screen "RIO 02 Digital Inputs" 1280x800, template "Template"
   on GenerateScreen: "TitleUpdater"()
   TextField "Text field_37" at 16,52 size 476x26; Text 'RIO #2 (Remote Inputs & Outputs Panel No. 2)'
   TextField "Text field_38" at 16,122 size 55x22; Text 'I15.0'
   TextField "Text field_39" at 16,157 size 55x22; Text 'I15.1'
   TextField "Text field_40" at 16,193 size 55x22; Text 'I15.2'
   TextField "Text field_41" at 16,229 size 55x22; Text 'I15.3'
   TextField "Text field_42" at 16,265 size 55x22; Text 'I15.4'
   TextField "Text field_43" at 16,301 size 55x22; Text 'I15.5'
   TextField "Text field_44" at 16,337 size 55x22; Text 'I15.6'
   TextField "Text field_45" at 16,373 size 55x22; Text 'I15.7'
   Circle "Circle_33" at 76,123 size 20x20
      Appearance <- "Tank 2P GTT Isolation Valve Feedback - Opened"
   Circle "Circle_34" at 76,158 size 20x20
      Appearance <- "Tank 2P GTT Isolation Valve Feedback - Closed"
   Circle "Circle_35" at 76,194 size 20x20
      Appearance <- "Tank 2P Tank Vent Valve 1 Feedback - Opened"
   Circle "Circle_36" at 76,230 size 20x20
      Appearance <- "Tank 2P Tank Vent Valve 1 Feedback - Closed"
   Circle "Circle_37" at 76,265 size 20x20
      Appearance <- "Tank 2P Tank Vent Valve 2 Feedback - Opened"
   Circle "Circle_38" at 76,301 size 20x20
      Appearance <- "Tank 2P Tank Vent Valve 2 Feedback - Closed"
   Circle "Circle_39" at 76,337 size 20x20
      Appearance <- "RIO2_SPR_DI_15_6"
   Circle "Circle_40" at 76,373 size 20x20
      Appearance <- "RIO2_SPR_DI_15_7"
   TextField "Text field_46" at 33,90 size 49x26; Text 'I0'
   TextField "Text field_47" at 16,441 size 55x22; Text 'I18.0'
   TextField "Text field_48" at 16,476 size 55x22; Text 'I18.1'
   TextField "Text field_49" at 16,512 size 55x22; Text 'I18.2'
   TextField "Text field_50" at 16,548 size 55x22; Text 'I18.3'
   TextField "Text field_51" at 16,584 size 55x22; Text 'I18.4'
   TextField "Text field_52" at 16,620 size 55x22; Text 'I18.5'
   TextField "Text field_53" at 16,656 size 55x22; Text 'I18.6'
   TextField "Text field_54" at 16,692 size 55x22; Text 'I18.7'
   Circle "Circle_41" at 76,442 size 20x20
      Appearance <- "Tank 2S GTT Isolation Valve Feedback - Opened"
   Circle "Circle_42" at 76,477 size 20x20
      Appearance <- "Tank 2S GTT Isolation Valve Feedback - Closed"
   Circle "Circle_43" at 76,513 size 20x20
      Appearance <- "Tank 2S Tank Vent Valve 1 Feedback - Opened"
   Circle "Circle_44" at 76,549 size 20x20
      Appearance <- "Tank 2S Tank Vent Valve 1 Feedback - Closed"
   Circle "Circle_45" at 76,585 size 20x20
      Appearance <- "Tank 2S Tank Vent Valve 2 Feedback - Opened"
   Circle "Circle_46" at 76,621 size 20x20
      Appearance <- "Tank 2S Tank Vent Valve 2 Feedback - Closed"
   Circle "Circle_47" at 76,657 size 20x20
      Appearance <- "RIO2_SPR_DI_18_6"
   Circle "Circle_48" at 76,693 size 20x20
      Appearance <- "RIO2_SPR_DI_18_7"
   TextField "Text field_55" at 33,409 size 49x26; Text 'I1'
   TextField "Text field_56" at 548,122 size 55x22; Text 'I21.0'
   TextField "Text field_57" at 548,157 size 55x22; Text 'I21.1'
   TextField "Text field_58" at 548,193 size 55x22; Text 'I21.2'
   TextField "Text field_59" at 548,229 size 55x22; Text 'I21.3'
   TextField "Text field_60" at 548,265 size 55x22; Text 'I21.4'
   TextField "Text field_61" at 548,301 size 55x22; Text 'I21.5'
   TextField "Text field_62" at 548,337 size 55x22; Text 'I21.6'
   TextField "Text field_63" at 548,373 size 55x22; Text 'I21.7'
   Circle "Circle_49" at 608,122 size 20x20
      Appearance <- "Tank 2P BWT Level High High Switch"
   Circle "Circle_50" at 608,157 size 20x20
      Appearance <- "RIO2 Tanks Pressure Switch Hi Hi"
   Circle "Circle_51" at 608,193 size 20x20
      Appearance <- "Tank 2S BWT Level High High Switch"
   Circle "Circle_52" at 608,229 size 20x20
      Appearance <- "RIO2_SPR_DI_21_3"
   Circle "Circle_53" at 608,265 size 20x20
      Appearance <- "RIO2_SPR_DI_21_4"
   Circle "Circle_54" at 608,301 size 20x20
      Appearance <- "RIO2_SPR_DI_21_5"
   Circle "Circle_55" at 608,337 size 20x20
      Appearance <- "RIO2_SPR_DI_21_6"
   Circle "Circle_56" at 608,373 size 20x20
      Appearance <- "RIO2_SPR_DI_21_7"
   TextField "Text field_64" at 570,90 size 49x26; Text 'I2'
   Button "HmiScreenItemData_1" at 1,1 size 150x43; TextOn 'Back'; TextOff 'Commissioning'
      on Release: ActivateScreen("Commissioning Main Page", 0)
   TextField "Text field_107" at 105,114 size 382x38; Text 'Tank 2P GTT Isolation Valve Feedback - Opened CV422'
   TextField "Text field_108" at 105,149 size 374x38; Text 'Tank 2P GTT Isolation Valve Feedback - Closed CV422'
   TextField "Text field_109" at 105,184 size 371x38; Text 'Tank 2P Tank Vent Valve 1 Feedback - Opened CV441-2P1'
   TextField "Text field_110" at 105,220 size 363x38; Text 'Tank 2P Tank Vent Valve 1 Feedback - Closed CV441-2P1'
   TextField "Text field_111" at 105,255 size 371x38; Text 'Tank 2P Tank Vent Valve 2 Feedback - Opened CV441-2P2'
   TextField "Text field_112" at 105,291 size 363x38; Text 'Tank 2P Tank Vent Valve 2 Feedback - Closed CV441-2P2'
   TextField "Text field_113" at 104,328 size 100x21; Text 'Spare Input'
   TextField "Text field_114" at 104,365 size 100x21; Text 'Spare Input'
   TextField "Text field_116" at 102,429 size 382x38; Text 'Tank 2S GTT Isolation Valve Feedback - Opened CV421-2S'
   TextField "Text field_117" at 102,465 size 374x38; Text 'Tank 2S GTT Isolation Valve Feedback - Closed CV421-2S'
   TextField "Text field_118" at 102,501 size 371x38; Text 'Tank 2S Tank Vent Valve 1 Feedback - Opened CV440-2SA'
   TextField "Text field_119" at 102,537 size 363x38; Text 'Tank 2S Tank Vent Valve 1 Feedback - Closed CV440-2SA'
   TextField "Text field_120" at 102,573 size 371x38; Text 'Tank 2S Tank Vent Valve 2 Feedback - Opened CV440-2SB'
   TextField "Text field_121" at 102,609 size 363x38; Text 'Tank 2S Tank Vent Valve 2 Feedback - Closed CV440-2SB'
   TextField "Text field_122" at 102,690 size 100x21; Text 'Spare Input'
   TextField "Text field_123" at 636,113 size 294x38; Text 'Tank 2P BWT Level High High Switch LS425-2P'
   TextField "Text field_124" at 636,148 size 270x38; Text 'RIO2 Tanks Pressure Switch Hi Hi PS436-2P/2S'
   TextField "Text field_125" at 636,184 size 294x38; Text 'Tank 2S BWT Level High High Switch LS422-2S'
   TextField "Text field_126" at 636,219 size 100x21; Text 'Spare Input'
   TextField "Text field_127" at 636,255 size 100x21; Text 'Spare Input'
   TextField "Text field_128" at 636,291 size 100x21; Text 'Spare Input'
   TextField "Text field_129" at 636,328 size 100x21; Text 'Spare Input'
   TextField "Text field_130" at 636,366 size 100x21; Text 'Spare Input'
   TextField "Text field_115" at 102,654 size 100x21; Text 'Spare Input'
   AlarmView "Alarm view_1" at 0,777 size 1280x23
   Group "Group" at 455,41 size 373x50
   Button "HmiScreenItemData_8" at 469,45 size 355x40; TextOn 'Back'; TextOff 'Text'
      on Click: "TitleUpdater"()
   TextField "Screen title" at 455,41 size 373x50; Text 'Screen title'

screen "RIO 03 Digital Inputs" 1280x800, template "Template"
   on GenerateScreen: "TitleUpdater"()
   TextField "Text field_37" at 16,52 size 476x26; Text 'RIO #3 (Remote Inputs & Outputs Panel No. 3)'
   TextField "Text field_38" at 16,122 size 55x22; Text 'I27.0'
   TextField "Text field_39" at 16,157 size 55x22; Text 'I27.1'
   TextField "Text field_40" at 16,193 size 55x22; Text 'I27.2'
   TextField "Text field_41" at 16,229 size 55x22; Text 'I27.3'
   TextField "Text field_42" at 16,265 size 55x22; Text 'I27.4'
   TextField "Text field_43" at 16,301 size 55x22; Text 'I27.5'
   TextField "Text field_44" at 16,337 size 55x22; Text 'I27.6'
   TextField "Text field_45" at 16,373 size 55x22; Text 'I27.7'
   Circle "Circle_33" at 76,123 size 20x20
      Appearance <- "Tank 3P GTT Isolation Valve Feedback - Opened"
   Circle "Circle_34" at 76,158 size 20x20
      Appearance <- "Tank 3P GTT Isolation Valve Feedback - Closed"
   Circle "Circle_35" at 76,194 size 20x20
      Appearance <- "Tank 3P Tank Vent Valve 1 Feedback - Opened"
   Circle "Circle_36" at 76,230 size 20x20
      Appearance <- "Tank 3P Tank Vent Valve 1 Feedback - Closed"
   Circle "Circle_37" at 76,265 size 20x20
      Appearance <- "Tank 3P Tank Vent Valve 2 Feedback - Opened"
   Circle "Circle_38" at 76,301 size 20x20
      Appearance <- "Tank 3P Tank Vent Valve 2 Feedback - Closed"
   Circle "Circle_39" at 76,337 size 20x20
      Appearance <- "RIO3_SPR_DI_27_6"
   Circle "Circle_40" at 76,373 size 20x20
      Appearance <- "RIO3_SPR_DI_27_7"
   TextField "Text field_46" at 33,90 size 49x26; Text 'I0'
   TextField "Text field_47" at 16,441 size 55x22; Text 'I30.0'
   TextField "Text field_48" at 16,476 size 55x22; Text 'I30.1'
   TextField "Text field_49" at 16,512 size 55x22; Text 'I30.2'
   TextField "Text field_50" at 16,548 size 55x22; Text 'I30.3'
   TextField "Text field_51" at 16,584 size 55x22; Text 'I30.4'
   TextField "Text field_52" at 16,620 size 55x22; Text 'I30.5'
   TextField "Text field_53" at 16,656 size 55x22; Text 'I30.6'
   TextField "Text field_54" at 16,692 size 55x22; Text 'I30.7'
   Circle "Circle_41" at 76,442 size 20x20
      Appearance <- "Tank 3S GTT Isolation Valve Feedback - Opened"
   Circle "Circle_42" at 76,477 size 20x20
      Appearance <- "Tank 3S GTT Isolation Valve Feedback - Closed"
   Circle "Circle_43" at 76,513 size 20x20
      Appearance <- "Tank 3S Tank Vent Valve 1 Feedback - Opened"
   Circle "Circle_44" at 76,549 size 20x20
      Appearance <- "Tank 3S Tank Vent Valve 1 Feedback - Closed"
   Circle "Circle_45" at 76,585 size 20x20
      Appearance <- "Tank 3S Tank Vent Valve 2 Feedback - Opened"
   Circle "Circle_46" at 76,621 size 20x20
      Appearance <- "Tank 3S Tank Vent Valve 2 Feedback - Closed"
   Circle "Circle_47" at 76,657 size 20x20
      Appearance <- "RIO3_SPR_DI_30_6"
   Circle "Circle_48" at 76,693 size 20x20
      Appearance <- "RIO3_SPR_DI_30_7"
   TextField "Text field_55" at 33,409 size 49x26; Text 'I1'
   TextField "Text field_56" at 548,122 size 55x22; Text 'I33.0'
   TextField "Text field_57" at 548,157 size 55x22; Text 'I33.1'
   TextField "Text field_58" at 548,193 size 55x22; Text 'I33.2'
   TextField "Text field_59" at 548,229 size 55x22; Text 'I33.3'
   TextField "Text field_60" at 548,265 size 55x22; Text 'I33.4'
   TextField "Text field_61" at 548,301 size 55x22; Text 'I33.5'
   TextField "Text field_62" at 548,337 size 55x22; Text 'I33.6'
   TextField "Text field_63" at 548,373 size 55x22; Text 'I33.7'
   Circle "Circle_49" at 608,122 size 20x20
      Appearance <- "Tank 3P BWT Level High High Switch"
   Circle "Circle_50" at 608,157 size 20x20
      Appearance <- "RIO3 Tanks Pressure Switch Hi Hi"
   Circle "Circle_51" at 608,193 size 20x20
      Appearance <- "Tank 3S BWT Level High High Switch"
   Circle "Circle_52" at 608,229 size 20x20
      Appearance <- "RIO3_SPR_DI_33_3"
   Circle "Circle_53" at 608,265 size 20x20
      Appearance <- "RIO3_SPR_DI_33_4"
   Circle "Circle_54" at 608,301 size 20x20
      Appearance <- "RIO3_SPR_DI_33_5"
   Circle "Circle_55" at 608,337 size 20x20
      Appearance <- "RIO3_SPR_DI_33_6"
   Circle "Circle_56" at 608,373 size 20x20
      Appearance <- "RIO3_SPR_DI_33_7"
   TextField "Text field_64" at 570,90 size 49x26; Text 'I2'
   Button "HmiScreenItemData_1" at 1,1 size 150x43; TextOn 'Back'; TextOff 'Commissioning'
      on Release: ActivateScreen("Commissioning Main Page", 0)
   TextField "Text field_107" at 105,114 size 382x38; Text 'Tank 3P GTT Isolation Valve Feedback - Opened CV422'
   TextField "Text field_108" at 105,149 size 374x38; Text 'Tank 3P GTT Isolation Valve Feedback - Closed CV422'
   TextField "Text field_109" at 105,184 size 371x38; Text 'Tank 3P Tank Vent Valve 1 Feedback - Opened CV441-3P1'
   TextField "Text field_110" at 105,220 size 363x38; Text 'Tank 3P Tank Vent Valve 1 Feedback - Closed CV441-3P1'
   TextField "Text field_111" at 105,255 size 371x38; Text 'Tank 3P Tank Vent Valve 2 Feedback - Opened CV441-3P2'
   TextField "Text field_112" at 105,291 size 363x38; Text 'Tank 3P Tank Vent Valve 2 Feedback - Closed CV441-3P2'
   TextField "Text field_113" at 104,328 size 100x21; Text 'Spare Input'
   TextField "Text field_114" at 104,365 size 100x21; Text 'Spare Input'
   TextField "Text field_116" at 102,429 size 382x38; Text 'Tank 3S GTT Isolation Valve Feedback - Opened CV421-3S'
   TextField "Text field_117" at 102,465 size 374x38; Text 'Tank 3S GTT Isolation Valve Feedback - Closed CV421-3S'
   TextField "Text field_118" at 102,501 size 371x38; Text 'Tank 3S Tank Vent Valve 1 Feedback - Opened CV440-3SA'
   TextField "Text field_119" at 102,537 size 363x38; Text 'Tank 3S Tank Vent Valve 1 Feedback - Closed CV440-3SA'
   TextField "Text field_120" at 102,573 size 371x38; Text 'Tank 3S Tank Vent Valve 2 Feedback - Opened CV440-3SB'
   TextField "Text field_121" at 102,609 size 363x38; Text 'Tank 3S Tank Vent Valve 2 Feedback - Closed CV440-3SB'
   TextField "Text field_122" at 102,690 size 100x21; Text 'Spare Input'
   TextField "Text field_123" at 636,113 size 294x38; Text 'Tank 3P BWT Level High High Switch LS425-3P'
   TextField "Text field_124" at 636,148 size 270x38; Text 'RIO3 Tanks Pressure Switch Hi Hi PS436-3P/3S'
   TextField "Text field_125" at 636,184 size 294x38; Text 'Tank 3S BWT Level High High Switch LS422-3S'
   TextField "Text field_126" at 636,219 size 100x21; Text 'Spare Input'
   TextField "Text field_127" at 636,255 size 100x21; Text 'Spare Input'
   TextField "Text field_128" at 636,291 size 100x21; Text 'Spare Input'
   TextField "Text field_129" at 636,328 size 100x21; Text 'Spare Input'
   TextField "Text field_130" at 636,366 size 100x21; Text 'Spare Input'
   TextField "Text field_115" at 102,654 size 100x21; Text 'Spare Input'
   AlarmView "Alarm view_1" at 0,777 size 1280x23
   Group "Group" at 455,41 size 373x50
   Button "HmiScreenItemData_8" at 469,45 size 355x40; TextOn 'Back'; TextOff 'Text'
      on Click: "TitleUpdater"()
   TextField "Screen title" at 455,41 size 373x50; Text 'Screen title'

screen "RIO 04 Digital Inputs" 1280x800, template "Template"
   on GenerateScreen: "TitleUpdater"()
   TextField "Text field_37" at 16,52 size 476x26; Text 'RIO #4 (Remote Inputs & Outputs Panel No. 4)'
   TextField "Text field_38" at 16,122 size 55x22; Text 'I39.0'
   TextField "Text field_39" at 16,157 size 55x22; Text 'I39.1'
   TextField "Text field_40" at 16,193 size 55x22; Text 'I39.2'
   TextField "Text field_41" at 16,229 size 55x22; Text 'I39.3'
   TextField "Text field_42" at 16,265 size 55x22; Text 'I39.4'
   TextField "Text field_43" at 16,301 size 55x22; Text 'I39.5'
   TextField "Text field_44" at 16,337 size 55x22; Text 'I39.6'
   TextField "Text field_45" at 16,373 size 55x22; Text 'I39.7'
   Circle "Circle_33" at 76,123 size 20x20
      Appearance <- "Tank 4P GTT Isolation Valve Feedback - Opened"
   Circle "Circle_34" at 76,158 size 20x20
      Appearance <- "Tank 4P GTT Isolation Valve Feedback - Closed"
   Circle "Circle_35" at 76,194 size 20x20
      Appearance <- "Tank 4P Tank Vent Valve 1 Feedback - Opened"
   Circle "Circle_36" at 76,230 size 20x20
      Appearance <- "Tank 4P Tank Vent Valve 1 Feedback - Closed"
   Circle "Circle_37" at 76,265 size 20x20
      Appearance <- "Tank 4P Tank Vent Valve 2 Feedback - Opened"
   Circle "Circle_38" at 76,301 size 20x20
      Appearance <- "Tank 4P Tank Vent Valve 2 Feedback - Closed"
   Circle "Circle_39" at 76,337 size 20x20
      Appearance <- "RIO4_SPR_DI_139_6"
   Circle "Circle_40" at 76,373 size 20x20
      Appearance <- "RIO4_SPR_DI_139_7"
   TextField "Text field_46" at 33,90 size 49x26; Text 'I0'
   TextField "Text field_47" at 16,441 size 55x22; Text 'I42.0'
   TextField "Text field_48" at 16,476 size 55x22; Text 'I42.1'
   TextField "Text field_49" at 16,512 size 55x22; Text 'I42.2'
   TextField "Text field_50" at 16,548 size 55x22; Text 'I42.3'
   TextField "Text field_51" at 16,584 size 55x22; Text 'I42.4'
   TextField "Text field_52" at 16,620 size 55x22; Text 'I42.5'
   TextField "Text field_53" at 16,656 size 55x22; Text 'I42.6'
   TextField "Text field_54" at 16,692 size 55x22; Text 'I42.7'
   Circle "Circle_41" at 76,442 size 20x20
      Appearance <- "Tank 4S GTT Isolation Valve Feedback - Opened"
   Circle "Circle_42" at 76,477 size 20x20
      Appearance <- "Tank 4S GTT Isolation Valve Feedback - Closed"
   Circle "Circle_43" at 76,513 size 20x20
      Appearance <- "Tank 4S Tank Vent Valve 1 Feedback - Opened"
   Circle "Circle_44" at 76,549 size 20x20
      Appearance <- "Tank 4S Tank Vent Valve 1 Feedback - Closed"
   Circle "Circle_45" at 76,585 size 20x20
      Appearance <- "Tank 4S Tank Vent Valve 2 Feedback - Opened"
   Circle "Circle_46" at 76,621 size 20x20
      Appearance <- "Tank 4S Tank Vent Valve 2 Feedback - Closed"
   Circle "Circle_47" at 76,657 size 20x20
      Appearance <- "RIO4_SPR_DI_142_6"
   Circle "Circle_48" at 76,693 size 20x20
      Appearance <- "RIO4_SPR_DI_142_7"
   TextField "Text field_55" at 33,409 size 49x26; Text 'I1'
   TextField "Text field_56" at 548,122 size 55x22; Text 'I45.0'
   TextField "Text field_57" at 548,157 size 55x22; Text 'I45.1'
   TextField "Text field_58" at 548,193 size 55x22; Text 'I45.2'
   TextField "Text field_59" at 548,229 size 55x22; Text 'I45.3'
   TextField "Text field_60" at 548,265 size 55x22; Text 'I45.4'
   TextField "Text field_61" at 548,301 size 55x22; Text 'I45.5'
   TextField "Text field_62" at 548,337 size 55x22; Text 'I45.6'
   TextField "Text field_63" at 548,373 size 55x22; Text 'I45.7'
   Circle "Circle_49" at 608,122 size 20x20
      Appearance <- "Tank 4P BWT Level High High Switch"
   Circle "Circle_50" at 608,157 size 20x20
      Appearance <- "RIO4 Tanks Pressure Switch Hi Hi"
   Circle "Circle_51" at 608,193 size 20x20
      Appearance <- "Tank 4S BWT Level High High Switch"
   Circle "Circle_52" at 608,229 size 20x20
      Appearance <- "RIO4_SPR_DI_145_3"
   Circle "Circle_53" at 608,265 size 20x20
      Appearance <- "RIO4_SPR_DI_145_4"
   Circle "Circle_54" at 608,301 size 20x20
      Appearance <- "RIO4_SPR_DI_145_5"
   Circle "Circle_55" at 608,337 size 20x20
      Appearance <- "RIO4_SPR_DI_145_6"
   Circle "Circle_56" at 608,373 size 20x20
      Appearance <- "RIO4_SPR_DI_145_7"
   TextField "Text field_64" at 570,90 size 49x26; Text 'I2'
   Button "HmiScreenItemData_1" at 1,1 size 150x43; TextOn 'Back'; TextOff 'Commissioning'
      on Release: ActivateScreen("Commissioning Main Page", 0)
   TextField "Text field_107" at 105,114 size 382x38; Text 'Tank 4P GTT Isolation Valve Feedback - Opened CV422'
   TextField "Text field_108" at 105,149 size 374x38; Text 'Tank 4P GTT Isolation Valve Feedback - Closed CV422'
   TextField "Text field_109" at 105,184 size 371x38; Text 'Tank 4P Tank Vent Valve 1 Feedback - Opened CV441-4P1'
   TextField "Text field_110" at 105,220 size 363x38; Text 'Tank 4P Tank Vent Valve 1 Feedback - Closed CV441-4P1'
   TextField "Text field_111" at 105,255 size 371x38; Text 'Tank 4P Tank Vent Valve 2 Feedback - Opened CV441-4P2'
   TextField "Text field_112" at 105,291 size 363x38; Text 'Tank 4P Tank Vent Valve 2 Feedback - Closed CV441-4P2'
   TextField "Text field_113" at 104,328 size 100x21; Text 'Spare Input'
   TextField "Text field_114" at 104,365 size 100x21; Text 'Spare Input'
   TextField "Text field_116" at 102,429 size 382x38; Text 'Tank 4S GTT Isolation Valve Feedback - Opened CV421-4S'
   TextField "Text field_117" at 102,465 size 374x38; Text 'Tank 4S GTT Isolation Valve Feedback - Closed CV421-4S'
   TextField "Text field_118" at 102,501 size 371x38; Text 'Tank 4S Tank Vent Valve 1 Feedback - Opened CV440-4SA'
   TextField "Text field_119" at 102,537 size 363x38; Text 'Tank 4S Tank Vent Valve 1 Feedback - Closed CV440-4SA'
   TextField "Text field_120" at 102,573 size 371x38; Text 'Tank 4S Tank Vent Valve 2 Feedback - Opened CV440-4SB'
   TextField "Text field_121" at 102,609 size 363x38; Text 'Tank 4S Tank Vent Valve 2 Feedback - Closed CV440-4SB'
   TextField "Text field_122" at 102,690 size 100x21; Text 'Spare Input'
   TextField "Text field_123" at 636,113 size 294x38; Text 'Tank 4P BWT Level High High Switch LS425-4P'
   TextField "Text field_124" at 636,148 size 270x38; Text 'RIO4 Tanks Pressure Switch Hi Hi PS436-4P/4S'
   TextField "Text field_125" at 636,184 size 294x38; Text 'Tank 3S BWT Level High High Switch LS422-4S'
   TextField "Text field_126" at 636,219 size 100x21; Text 'Spare Input'
   TextField "Text field_127" at 636,255 size 100x21; Text 'Spare Input'
   TextField "Text field_128" at 636,291 size 100x21; Text 'Spare Input'
   TextField "Text field_129" at 636,328 size 100x21; Text 'Spare Input'
   TextField "Text field_130" at 636,366 size 100x21; Text 'Spare Input'
   TextField "Text field_115" at 102,654 size 100x21; Text 'Spare Input'
   AlarmView "Alarm view_1" at 0,777 size 1280x23
   Group "Group" at 455,41 size 373x50
   Button "HmiScreenItemData_8" at 469,45 size 355x40; TextOn 'Back'; TextOff 'Text'
      on Click: "TitleUpdater"()
   TextField "Screen title" at 455,41 size 373x50; Text 'Screen title'

screen "RIO 05 Digital Inputs" 1280x800, template "Template"
   on GenerateScreen: "TitleUpdater"()
   TextField "Text field_37" at 16,52 size 476x26; Text 'RIO #5 (Remote Inputs & Outputs Panel No. 5)'
   TextField "Text field_38" at 16,122 size 55x22; Text 'I51.0'
   TextField "Text field_39" at 16,157 size 55x22; Text 'I51.1'
   TextField "Text field_40" at 16,193 size 55x22; Text 'I51.2'
   TextField "Text field_41" at 16,229 size 55x22; Text 'I51.3'
   TextField "Text field_42" at 16,265 size 55x22; Text 'I51.4'
   TextField "Text field_43" at 16,301 size 55x22; Text 'I51.5'
   TextField "Text field_44" at 16,337 size 55x22; Text 'I51.6'
   TextField "Text field_45" at 16,373 size 55x22; Text 'I51.7'
   Circle "Circle_33" at 76,123 size 20x20
      Appearance <- "Tank 5P GTT Isolation Valve Feedback - Opened"
   Circle "Circle_34" at 76,158 size 20x20
      Appearance <- "Tank 5P GTT Isolation Valve Feedback - Closed"
   Circle "Circle_35" at 76,194 size 20x20
      Appearance <- "Tank 5P Tank Vent Valve 1 Feedback - Opened"
   Circle "Circle_36" at 76,230 size 20x20
      Appearance <- "Tank 5P Tank Vent Valve 1 Feedback - Closed"
   Circle "Circle_37" at 76,265 size 20x20
      Appearance <- "Tank 5P Tank Vent Valve 2 Feedback - Opened"
   Circle "Circle_38" at 76,301 size 20x20
      Appearance <- "Tank 5P Tank Vent Valve 2 Feedback - Closed"
   Circle "Circle_39" at 76,337 size 20x20
      Appearance <- "RIO5_SPR_DI_51_6"
   Circle "Circle_40" at 76,373 size 20x20
      Appearance <- "RIO5_SPR_DI_51_7"
   TextField "Text field_46" at 33,90 size 49x26; Text 'I0'
   TextField "Text field_47" at 16,441 size 55x22; Text 'I54.0'
   TextField "Text field_48" at 16,476 size 55x22; Text 'I54.1'
   TextField "Text field_49" at 16,512 size 55x22; Text 'I54.2'
   TextField "Text field_50" at 16,548 size 55x22; Text 'I54.3'
   TextField "Text field_51" at 16,584 size 55x22; Text 'I54.4'
   TextField "Text field_52" at 16,620 size 55x22; Text 'I54.5'
   TextField "Text field_53" at 16,656 size 55x22; Text 'I54.6'
   TextField "Text field_54" at 16,692 size 55x22; Text 'I54.7'
   Circle "Circle_41" at 76,442 size 20x20
      Appearance <- "Tank 5S GTT Isolation Valve Feedback - Opened"
   Circle "Circle_42" at 76,477 size 20x20
      Appearance <- "Tank 5S GTT Isolation Valve Feedback - Closed"
   Circle "Circle_43" at 76,513 size 20x20
      Appearance <- "Tank 5S Tank Vent Valve 1 Feedback - Opened"
   Circle "Circle_44" at 76,549 size 20x20
      Appearance <- "Tank 5S Tank Vent Valve 1 Feedback - Closed"
   Circle "Circle_45" at 76,585 size 20x20
      Appearance <- "Tank 5S Tank Vent Valve 2 Feedback - Opened"
   Circle "Circle_46" at 76,621 size 20x20
      Appearance <- "Tank 5S Tank Vent Valve 2 Feedback - Closed"
   Circle "Circle_47" at 76,657 size 20x20
      Appearance <- "RIO5_SPR_DI_54_6"
   Circle "Circle_48" at 76,693 size 20x20
      Appearance <- "RIO5_SPR_DI_54_7"
   TextField "Text field_55" at 33,409 size 49x26; Text 'I1'
   TextField "Text field_56" at 548,122 size 55x22; Text 'I57.0'
   TextField "Text field_57" at 548,157 size 55x22; Text 'I57.1'
   TextField "Text field_58" at 548,193 size 55x22; Text 'I57.2'
   TextField "Text field_59" at 548,229 size 55x22; Text 'I57.3'
   TextField "Text field_60" at 548,265 size 55x22; Text 'I57.4'
   TextField "Text field_61" at 548,301 size 55x22; Text 'I57.5'
   TextField "Text field_62" at 548,337 size 55x22; Text 'I57.6'
   TextField "Text field_63" at 548,373 size 55x22; Text 'I57.7'
   Circle "Circle_49" at 608,122 size 20x20
      Appearance <- "Tank 5P BWT Level High High Switch"
   Circle "Circle_50" at 608,157 size 20x20
      Appearance <- "RIO5 Tanks Pressure Switch Hi Hi"
   Circle "Circle_51" at 608,193 size 20x20
      Appearance <- "Tank 5S BWT Level High High Switch"
   Circle "Circle_52" at 608,229 size 20x20
      Appearance <- "RIO5_SPR_DI_57_3"
   Circle "Circle_53" at 608,265 size 20x20
      Appearance <- "RIO5_SPR_DI_57_4"
   Circle "Circle_54" at 608,301 size 20x20
      Appearance <- "RIO5_SPR_DI_57_5"
   Circle "Circle_55" at 608,337 size 20x20
      Appearance <- "RIO5_SPR_DI_57_6"
   Circle "Circle_56" at 608,373 size 20x20
      Appearance <- "RIO5_SPR_DI_57_7"
   TextField "Text field_64" at 570,90 size 49x26; Text 'I2'
   Button "HmiScreenItemData_1" at 1,1 size 150x43; TextOn 'Back'; TextOff 'Commissioning'
      on Release: ActivateScreen("Commissioning Main Page", 0)
   TextField "Text field_107" at 105,114 size 382x38; Text 'Tank 5P GTT Isolation Valve Feedback - Opened CV422'
   TextField "Text field_108" at 105,149 size 374x38; Text 'Tank 5P GTT Isolation Valve Feedback - Closed CV422'
   TextField "Text field_109" at 105,184 size 371x38; Text 'Tank 5P Tank Vent Valve 1 Feedback - Opened CV441-5P1'
   TextField "Text field_110" at 105,220 size 363x38; Text 'Tank 5P Tank Vent Valve 1 Feedback - Closed CV441-5P1'
   TextField "Text field_111" at 105,255 size 371x38; Text 'Tank 5P Tank Vent Valve 2 Feedback - Opened CV441-5P2'
   TextField "Text field_112" at 105,291 size 363x38; Text 'Tank 5P Tank Vent Valve 2 Feedback - Closed CV441-5P2'
   TextField "Text field_113" at 104,328 size 100x21; Text 'Spare Input'
   TextField "Text field_114" at 104,365 size 100x21; Text 'Spare Input'
   TextField "Text field_116" at 102,429 size 382x38; Text 'Tank 5S GTT Isolation Valve Feedback - Opened CV421-5S'
   TextField "Text field_117" at 102,465 size 374x38; Text 'Tank 5S GTT Isolation Valve Feedback - Closed CV421-5S'
   TextField "Text field_118" at 102,501 size 371x38; Text 'Tank 5S Tank Vent Valve 1 Feedback - Opened CV440-5SA'
   TextField "Text field_119" at 102,537 size 363x38; Text 'Tank 5S Tank Vent Valve 1 Feedback - Closed CV440-5SA'
   TextField "Text field_120" at 102,573 size 371x38; Text 'Tank 5S Tank Vent Valve 2 Feedback - Opened CV440-5SB'
   TextField "Text field_121" at 102,609 size 363x38; Text 'Tank 5S Tank Vent Valve 2 Feedback - Closed CV440-5SB'
   TextField "Text field_122" at 102,690 size 100x21; Text 'Spare Input'
   TextField "Text field_123" at 636,113 size 294x38; Text 'Tank 5P BWT Level High High Switch LS425-5P'
   TextField "Text field_124" at 636,148 size 270x38; Text 'RIO5 Tanks Pressure Switch Hi Hi PS436-5P/5S'
   TextField "Text field_125" at 636,184 size 294x38; Text 'Tank 5S BWT Level High High Switch LS422-5S'
   TextField "Text field_126" at 636,219 size 100x21; Text 'Spare Input'
   TextField "Text field_127" at 636,255 size 100x21; Text 'Spare Input'
   TextField "Text field_128" at 636,291 size 100x21; Text 'Spare Input'
   TextField "Text field_129" at 636,328 size 100x21; Text 'Spare Input'
   TextField "Text field_130" at 636,366 size 100x21; Text 'Spare Input'
   TextField "Text field_115" at 102,654 size 100x21; Text 'Spare Input'
   AlarmView "Alarm view_1" at 0,777 size 1280x23
   Group "Group" at 455,41 size 373x50
   Button "HmiScreenItemData_8" at 469,45 size 355x40; TextOn 'Back'; TextOff 'Text'
      on Click: "TitleUpdater"()
   TextField "Screen title" at 455,41 size 373x50; Text 'Screen title'

screen "RIO 06 Digital Inputs" 1280x800, template "Template"
   on GenerateScreen: "TitleUpdater"()
   TextField "Text field_37" at 16,52 size 476x26; Text 'RIO #6 (Remote Inputs & Outputs Panel No. 6)'
   TextField "Text field_38" at 16,122 size 55x22; Text 'I60.0'
   TextField "Text field_39" at 16,157 size 55x22; Text 'I60.1'
   TextField "Text field_40" at 16,193 size 55x22; Text 'I60.2'
   TextField "Text field_41" at 16,229 size 55x22; Text 'I60.3'
   TextField "Text field_42" at 16,265 size 55x22; Text 'I60.4'
   TextField "Text field_43" at 16,301 size 55x22; Text 'I60.5'
   TextField "Text field_44" at 16,337 size 55x22; Text 'I60.6'
   TextField "Text field_45" at 16,373 size 55x22; Text 'I60.7'
   Circle "Circle_33" at 76,123 size 20x20
      Appearance <- "Tank 6P GTT Isolation Valve Feedback - Opened"
   Circle "Circle_34" at 76,158 size 20x20
      Appearance <- "Tank 6P GTT Isolation Valve Feedback - Closed"
   Circle "Circle_35" at 76,194 size 20x20
      Appearance <- "Tank 6P Tank Vent Valve 1 Feedback - Opened"
   Circle "Circle_36" at 76,230 size 20x20
      Appearance <- "Tank 6P Tank Vent Valve 1 Feedback - Closed"
   Circle "Circle_37" at 76,265 size 20x20
      Appearance <- "Tank 6P Tank Vent Valve 2 Feedback - Opened"
   Circle "Circle_38" at 76,301 size 20x20
      Appearance <- "Tank 6P Tank Vent Valve 2 Feedback - Closed"
   Circle "Circle_39" at 76,337 size 20x20
      Appearance <- "RIO6_SPR_DI_60_6"
   Circle "Circle_40" at 76,373 size 20x20
      Appearance <- "RIO6_SPR_DI_60_7"
   TextField "Text field_46" at 33,90 size 49x26; Text 'I0'
   TextField "Text field_47" at 16,441 size 55x22; Text 'I63.0'
   TextField "Text field_48" at 16,476 size 55x22; Text 'I63.1'
   TextField "Text field_49" at 16,512 size 55x22; Text 'I63.2'
   TextField "Text field_50" at 16,548 size 55x22; Text 'I63.3'
   TextField "Text field_51" at 16,584 size 55x22; Text 'I63.4'
   TextField "Text field_52" at 16,620 size 55x22; Text 'I63.5'
   TextField "Text field_53" at 16,656 size 55x22; Text 'I63.6'
   TextField "Text field_54" at 16,692 size 55x22; Text 'I63.7'
   Circle "Circle_41" at 76,442 size 20x20
      Appearance <- "Tank 6S GTT Isolation Valve Feedback - Opened"
   Circle "Circle_42" at 76,477 size 20x20
      Appearance <- "Tank 6S GTT Isolation Valve Feedback - Closed"
   Circle "Circle_43" at 76,513 size 20x20
      Appearance <- "Tank 6S Tank Vent Valve 1 Feedback - Opened"
   Circle "Circle_44" at 76,549 size 20x20
      Appearance <- "Tank 6S Tank Vent Valve 1 Feedback - Closed"
   Circle "Circle_45" at 76,585 size 20x20
      Appearance <- "Tank 6S Tank Vent Valve 2 Feedback - Opened"
   Circle "Circle_46" at 76,621 size 20x20
      Appearance <- "Tank 6S Tank Vent Valve 2 Feedback - Closed"
   Circle "Circle_47" at 76,657 size 20x20
      Appearance <- "RIO6_SPR_DI_63_6"
   Circle "Circle_48" at 76,693 size 20x20
      Appearance <- "RIO6_SPR_DI_63_7"
   TextField "Text field_55" at 33,409 size 49x26; Text 'I1'
   TextField "Text field_56" at 548,122 size 55x22; Text 'I66.0'
   TextField "Text field_57" at 548,157 size 55x22; Text 'I66.1'
   TextField "Text field_58" at 548,193 size 55x22; Text 'I66.2'
   TextField "Text field_59" at 548,229 size 55x22; Text 'I66.3'
   TextField "Text field_60" at 548,265 size 55x22; Text 'I66.4'
   TextField "Text field_61" at 548,301 size 55x22; Text 'I66.5'
   TextField "Text field_62" at 548,337 size 55x22; Text 'I66.6'
   TextField "Text field_63" at 548,373 size 55x22; Text 'I66.7'
   Circle "Circle_49" at 608,122 size 20x20
      Appearance <- "Tank 6P BWT Level High High Switch"
   Circle "Circle_50" at 608,157 size 20x20
      Appearance <- "RIO6 Tanks Pressure Switch Hi Hi"
   Circle "Circle_51" at 608,193 size 20x20
      Appearance <- "Tank 6S BWT Level High High Switch"
   Circle "Circle_52" at 608,229 size 20x20
      Appearance <- "RIO6_SPR_DI_66_3"
   Circle "Circle_53" at 608,265 size 20x20
      Appearance <- "RIO6_SPR_DI_66_4"
   Circle "Circle_54" at 608,301 size 20x20
      Appearance <- "RIO6_SPR_DI_66_5"
   Circle "Circle_55" at 608,337 size 20x20
      Appearance <- "RIO6_SPR_DI_66_6"
   Circle "Circle_56" at 608,373 size 20x20
      Appearance <- "RIO6_SPR_DI_66_7"
   TextField "Text field_64" at 570,90 size 49x26; Text 'I2'
   Button "HmiScreenItemData_1" at 1,1 size 150x43; TextOn 'Back'; TextOff 'Commissioning'
      on Release: ActivateScreen("Commissioning Main Page", 0)
   TextField "Text field_107" at 105,114 size 382x38; Text 'Tank 6P GTT Isolation Valve Feedback - Opened CV422'
   TextField "Text field_108" at 105,149 size 374x38; Text 'Tank 6P GTT Isolation Valve Feedback - Closed CV422'
   TextField "Text field_109" at 105,184 size 371x38; Text 'Tank 6P Tank Vent Valve 1 Feedback - Opened CV441-6P1'
   TextField "Text field_110" at 105,220 size 363x38; Text 'Tank 6P Tank Vent Valve 1 Feedback - Closed CV441-6P1'
   TextField "Text field_111" at 105,255 size 371x38; Text 'Tank 6P Tank Vent Valve 2 Feedback - Opened CV441-6P2'
   TextField "Text field_112" at 105,291 size 363x38; Text 'Tank 6P Tank Vent Valve 2 Feedback - Closed CV441-6P2'
   TextField "Text field_113" at 104,328 size 100x21; Text 'Spare Input'
   TextField "Text field_114" at 104,365 size 100x21; Text 'Spare Input'
   TextField "Text field_116" at 102,429 size 382x38; Text 'Tank 6S GTT Isolation Valve Feedback - Opened CV421-6S'
   TextField "Text field_117" at 102,465 size 374x38; Text 'Tank 6S GTT Isolation Valve Feedback - Closed CV421-6S'
   TextField "Text field_118" at 102,501 size 371x38; Text 'Tank 6S Tank Vent Valve 1 Feedback - Opened CV440-6SA'
   TextField "Text field_119" at 102,537 size 363x38; Text 'Tank 6S Tank Vent Valve 1 Feedback - Closed CV440-6SA'
   TextField "Text field_120" at 102,573 size 371x38; Text 'Tank 6S Tank Vent Valve 2 Feedback - Opened CV440-6SB'
   TextField "Text field_121" at 102,609 size 363x38; Text 'Tank 6S Tank Vent Valve 2 Feedback - Closed CV440-6SB'
   TextField "Text field_122" at 102,690 size 100x21; Text 'Spare Input'
   TextField "Text field_123" at 636,113 size 294x38; Text 'Tank 6P BWT Level High High Switch LS425-6P'
   TextField "Text field_124" at 636,148 size 270x38; Text 'RIO6 Tanks Pressure Switch Hi Hi PS436-6P/6S'
   TextField "Text field_125" at 636,184 size 294x38; Text 'Tank 6S BWT Level High High Switch LS422-6S'
   TextField "Text field_126" at 636,219 size 100x21; Text 'Spare Input'
   TextField "Text field_127" at 636,255 size 100x21; Text 'Spare Input'
   TextField "Text field_128" at 636,291 size 100x21; Text 'Spare Input'
   TextField "Text field_129" at 636,328 size 100x21; Text 'Spare Input'
   TextField "Text field_130" at 636,366 size 100x21; Text 'Spare Input'
   TextField "Text field_115" at 102,654 size 100x21; Text 'Spare Input'
   AlarmView "Alarm view_1" at 0,777 size 1280x23
   Group "Group" at 455,41 size 373x50
   Button "HmiScreenItemData_8" at 469,45 size 355x40; TextOn 'Back'; TextOff 'Text'
      on Click: "TitleUpdater"()
   TextField "Screen title" at 455,41 size 373x50; Text 'Screen title'

screen "RIO 07 Digital Inputs" 1280x800, template "Template"
   on GenerateScreen: "TitleUpdater"()
   TextField "Text field_37" at 16,52 size 476x26; Text 'RIO #7 (Remote Inputs & Outputs Panel No. 7)'
   TextField "Text field_38" at 16,122 size 55x22; Text 'I75.0'
   TextField "Text field_39" at 16,157 size 55x22; Text 'I75.1'
   TextField "Text field_40" at 16,193 size 55x22; Text 'I75.2'
   TextField "Text field_41" at 16,229 size 55x22; Text 'I75.3'
   TextField "Text field_42" at 16,265 size 55x22; Text 'I75.4'
   TextField "Text field_43" at 16,301 size 55x22; Text 'I75.5'
   TextField "Text field_44" at 16,337 size 55x22; Text 'I75.6'
   TextField "Text field_45" at 16,373 size 55x22; Text 'I75.7'
   Circle "Circle_33" at 76,123 size 20x20
      Appearance <- "APT GTT Isolation Valve Feedback - Opened"
   Circle "Circle_34" at 76,158 size 20x20
      Appearance <- "APT GTT Isolation Valve Feedback - Closed"
   Circle "Circle_35" at 76,194 size 20x20
      Appearance <- "APT Tank Vent Valve 1 Feedback - Opened"
   Circle "Circle_36" at 76,230 size 20x20
      Appearance <- "APT Tank Vent Valve 1 Feedback - Closed"
   Circle "Circle_37" at 76,265 size 20x20
      Appearance <- "APT Tank Vent Valve 2 Feedback - Opened"
   Circle "Circle_38" at 76,301 size 20x20
      Appearance <- "APT Tank Vent Valve 2 Feedback - Closed"
   Circle "Circle_39" at 76,337 size 20x20
      Appearance <- "RIO7_SPR_DI_175_6"
   Circle "Circle_40" at 76,373 size 20x20
      Appearance <- "RIO7_SPR_DI_175_7"
   TextField "Text field_46" at 33,90 size 49x26; Text 'I0'
   TextField "Text field_56" at 548,122 size 55x22; Text 'I78.0'
   TextField "Text field_57" at 548,157 size 55x22; Text 'I78.1'
   TextField "Text field_58" at 548,193 size 55x22; Text 'I78.2'
   TextField "Text field_59" at 548,229 size 55x22; Text 'I78.3'
   TextField "Text field_60" at 548,265 size 55x22; Text 'I78.4'
   TextField "Text field_61" at 548,301 size 55x22; Text 'I78.5'
   TextField "Text field_62" at 548,337 size 55x22; Text 'I78.6'
   TextField "Text field_63" at 548,373 size 55x22; Text 'I78.7'
   Circle "Circle_49" at 608,122 size 20x20
      Appearance <- "APT BWT Level High High Switch"
   Circle "Circle_50" at 608,157 size 20x20
      Appearance <- "RIO7 Tank Pressure Switch Hi Hi"
   Circle "Circle_51" at 608,193 size 20x20
      Appearance <- "RIO7_SPR_DI_178_2"
   Circle "Circle_52" at 608,229 size 20x20
      Appearance <- "RIO7_SPR_DI_178_3"
   Circle "Circle_53" at 608,265 size 20x20
      Appearance <- "RIO7_SPR_DI_178_4"
   Circle "Circle_54" at 608,301 size 20x20
      Appearance <- "RIO7_SPR_DI_178_5"
   Circle "Circle_55" at 608,337 size 20x20
      Appearance <- "RIO7_SPR_DI_178_6"
   Circle "Circle_56" at 608,373 size 20x20
      Appearance <- "RIO7_SPR_DI_178_7"
   TextField "Text field_64" at 570,90 size 49x26; Text 'I1'
   Button "HmiScreenItemData_1" at 1,1 size 150x43; TextOn 'Back'; TextOff 'Commissioning'
      on Release: ActivateScreen("Commissioning Main Page", 0)
   TextField "Text field_107" at 105,114 size 393x38; Text 'Tank APT GTT Isolation Valve Feedback - Opened CV422'
   TextField "Text field_108" at 105,149 size 385x38; Text 'Tank APT GTT Isolation Valve Feedback - Closed CV422'
   TextField "Text field_109" at 105,184 size 382x38; Text 'Tank APT Tank Vent Valve 1 Feedback - Opened CV441-APT1'
   TextField "Text field_110" at 105,220 size 374x38; Text 'Tank APT Tank Vent Valve 1 Feedback - Closed CV441-APT1'
   TextField "Text field_111" at 105,255 size 382x38; Text 'Tank APT Tank Vent Valve 2 Feedback - Opened CV441-APT2'
   TextField "Text field_112" at 105,291 size 374x38; Text 'Tank APT Tank Vent Valve 2 Feedback - Closed CV441-APT2'
   TextField "Text field_113" at 104,328 size 100x21; Text 'Spare Input'
   TextField "Text field_114" at 104,365 size 100x21; Text 'Spare Input'
   TextField "Text field_123" at 636,113 size 294x38; Text 'Tank APT BWT Level High High Switch LS425-APT'
   TextField "Text field_124" at 636,148 size 270x38; Text 'RIO7 Tanks Pressure Switch Hi Hi PS436-APT'
   TextField "Text field_125" at 636,184 size 100x21; Text 'Spare Input'
   TextField "Text field_126" at 636,219 size 100x21; Text 'Spare Input'
   TextField "Text field_127" at 636,255 size 100x21; Text 'Spare Input'
   TextField "Text field_128" at 636,291 size 100x21; Text 'Spare Input'
   TextField "Text field_129" at 636,328 size 100x21; Text 'Spare Input'
   TextField "Text field_130" at 636,366 size 100x21; Text 'Spare Input'
   AlarmView "Alarm view_1" at 0,777 size 1280x23
   Group "Group" at 455,41 size 373x50
   Button "HmiScreenItemData_8" at 469,45 size 355x40; TextOn 'Back'; TextOff 'Text'
      on Click: "TitleUpdater"()
   TextField "Screen title" at 455,41 size 373x50; Text 'Screen title'

screen "04 Alarm Log" 1280x800, template "Template"
   AlarmView "Alarm view_1" at 8,61 size 1258x665
   Button "HmiScreenItemData_1" at 1,1 size 139x43; TextOn 'Back'; TextOff 'Main Index'
      on Release: ActivateScreen("02 Main Index", 0)
   Button "HmiScreenItemData_2" at 143,1 size 139x43; TextOn 'Back'; TextOff 'Alarm Buffer'
      on Release: ActivateScreen("05 Alarm Buffer", 0)
   Button "HmiScreenItemData_3" at 1124,735 size 139x43; TextOn 'RESET ALARMS'; TextOff 'Reset Alarms'
      on Click: function_d9204949("Alarm view_1")
      on Press: function_b14e0dd5("80_From_HMI_Reset_Alarms", 0)
   Button "HmiScreenItemData_18" at 953,735 size 139x43; TextOn 'Back'; TextOff 'Silence Buzzer'; Authorization "User administration"
      on Press: function_b14e0dd5("80_From_HMI_SLNCE_BZR", 0)
      Appearance <- "80_From_HMI_SLNCE_BZR"
   Button "HmiScreenItemData_4" at 1138,1 size 139x43; TextOn 'I&A Compressor Ok'; TextOff 'Back'
      on Release: function_efd93a16()

screen "Air System" 1280x800, template "Template"
   Button "Button_16" at 609,168 size 64x25; TextOn 'Alarm'; TextOff 'Text'
   Button "Button_2" at 602,168 size 71x25; TextOn 'Alarm'; TextOff 'Shutdown'
      Visibility <- "10 DI_DATA_E131_SHTDN"
   Button "HmiScreenItemData_1" at 1,1 size 150x43; TextOn 'Back'; TextOff 'Main Index'
      on Release: ActivateScreen("02 Main Index", 0)
   Button "Button_15" at 464,168 size 57x25; TextOn 'Enabled'; TextOff 'Disabled'
   TextField "Text field_14" at 307,171 size 158x18; Text 'I & A Air Compressor'
   TextField "Text field_15" at 464,146 size 60x18; Text 'Enabled'
   TextField "Text field_16" at 530,146 size 64x18; Text 'Running'
   TextField "Text field_18" at 601,145 size 78x18; Text 'Shutdown'
   Button "Button_1" at 530,168 size 57x25; TextOn 'Enabled'; TextOff 'Stopped'
   TextField "Text field_1" at 282,55 size 561x26; Text 'Instrument & Atomising Air Compressor Control (E-131)'
   TextField "Text field_32" at 464,168 size 57x25; Text 'Enabled'
      Visibility <- "14_DQ_Data_E131ControlOut"
   TextField "Text field_2" at 530,168 size 57x25; Text 'Running'
      Visibility <- "10 DI_DATA_E131_OK"
   GraphicIOField "Graphic I/O field_2" at 703,308 size 196x199; PictureList "IA Compressor_2"
      ProcessValue <- "82_To_HMI_CA Blower Animation"
   Gauge "Gauge_1" at 791,570 size 184x184; CaptionText 'Open'; UnitText '%'
      ProcessValue <- "12_AI_Data_CV403_SCALED"
   TextField "Text field_20" at 374,532 size 529x26; Text 'Combustion Air/Inert Gas Pressure Control (CV-403)'
   IOField "I/O field_16" at 516,441 size 74x25; FormatPattern 9999; Unit  RPM
      ProcessValue <- "12_AI_Data_E139_RPM_SCALED"
   IOField "I/O field_1" at 602,441 size 69x25; FormatPattern 999.99; Unit  A
      ProcessValue <- "12_AI_Data_E139_AMPS_SCALED"
   TextField "Text field_7" at 364,279 size 391x26; Text 'Combustion Air Blower Control (E-139)'
   Button "Button_3" at 464,395 size 57x25; TextOn 'Enabled'; TextOff 'Disabled'
   TextField "Text field_4" at 464,373 size 60x18; Text 'Enabled'
   TextField "Text field_5" at 624,373 size 40x18; Text 'Fault'
   Button "Button_5" at 615,396 size 57x25; TextOn 'Enabled'; TextOff 'Healthy'
   TextField "Text field_8" at 464,395 size 57x25; Text 'Enabled'
      Visibility <- "14_DQ_Data_E139_CNTRL"
   Button "Button_6" at 616,395 size 57x25; TextOn 'Alarm'; TextOff 'Fault'
      Visibility <- "10_DI_Data_E139_VSD_FLT"
      Appearance <- "10_DI_Data_E139_VSD_FLT"
   TextField "Text field_11" at 320,444 size 84x18; Text 'Motor RPM'
   TextField "Text field_3" at 307,399 size 124x18; Text 'Combustion Air'
   IOField "I/O field_5" at 429,441 size 75x25; Authorization "Operating Mode"; FormatPattern 9999; Unit  RPM
      ProcessValue <- "80_From_HMI_E139_SET_SPEED"
   Button "HmiScreenItemData_11" at 1016,173 size 69x51; TextOn 'RESET'; TextOff 'Reset'; Authorization "Operate"
      on Press: function_b14e0dd5("82_To_HMI_I&A Compressor Reset Hours", 0)
   IOField "I/O field_8" at 941,175 size 65x25; FormatPattern 99999; Unit  h
      ProcessValue <- "82_To_HMI_I&A Compressor Run Hours(1)"
   IOField "I/O field_9" at 941,205 size 65x25; Authorization "Operate"; FormatPattern 99999; Unit  h
      ProcessValue <- "82_To_HMI_I&A Compressor Service Time Hours"
   TextField "Text field_19" at 911,174 size 37x20; Text 'Run'
   TextField "Text field_21" at 911,205 size 37x20; Text 'Set'
   TextField "Text field_13" at 954,78 size 140x20; Text 'Service Hour E131'
   Button "HmiScreenItemData_12" at 1016,428 size 69x51; TextOn 'RESET'; TextOff 'Reset'; Authorization "Operate"
      on Press: function_b14e0dd5("82_To_HMI_CA Blower Reset Hours", 0)
   IOField "I/O field_10" at 941,427 size 65x25; FormatPattern 9999; Unit h
      ProcessValue <- "82_To_HMI_CA Blower Run Hours"
   IOField "I/O field_11" at 941,457 size 65x25; Authorization "Operate"; FormatPattern 9999; Unit  h
      ProcessValue <- "82_To_HMI_CA Blower Service Time Hours"
   TextField "Text field_22" at 911,429 size 37x20; Text 'Run'
   TextField "Text field_23" at 911,459 size 37x20; Text 'Set'
   TextField "Text field_24" at 954,329 size 148x20; Text 'Service Hours E139'
   Button "HmiScreenItemData_13" at 933,357 size 183x34; TextOn 'Back'; TextOff 'Text'
   IOField "I/O field_13" at 983,362 size 40x25; FormatPattern 99; Unit h
      ProcessValue <- "82_To_HMI_CA Blower Run Hours"
   IOField "I/O field_14" at 1025,362 size 40x25; FormatPattern 99; Unit m
      ProcessValue <- "82_To_HMI_CA Blower Run Minutes"
   IOField "I/O field_15" at 940,362 size 40x25; FormatPattern 99; Unit d
      ProcessValue <- "82_To_HMI_CA Blower Run Days"
   Button "HmiScreenItemData_14" at 928,105 size 183x34; TextOn 'Back'; TextOff 'Text'
   IOField "I/O field_17" at 978,109 size 40x25; FormatPattern 99; Unit h
      ProcessValue <- "82_To_HMI_I&A Compressor Run Hours"
   IOField "I/O field_18" at 1021,109 size 40x25; FormatPattern 99; Unit m
      ProcessValue <- "82_To_HMI_I&A Compressor Run Minutes"
   IOField "I/O field_19" at 1064,109 size 40x25; FormatPattern 99; Unit s
      ProcessValue <- "82_To_HMI_I&A Compressor Run Seconds"
   Button "Button_4" at 840,56 size 57x25; TextOn 'Alarm'; TextOff 'Service'
      Visibility <- "82_To_HMI_I&A Compressor Service Due"
   Button "Button_7" at 840,280 size 57x25; TextOn 'Alarm'; TextOff 'Service'
      Visibility <- "82_To_HMI_CA Blower Service Due"
   TextField "Text field_26" at 773,754 size 224x22; Text 'Modulating Valve Position'
   GraphicView "Graphic view_91" at 713,108 size 113x127; Picture "Graphic_246"
   GraphicIOField "Graphic I/O field_5" at 705,101 size 128x139; PictureList "New IA Compressor"
      Visibility <- "68_Sys_Status_Data_IA_PRES_IN_RNG(1)"
      ProcessValue <- "82_To_HMI_IA Compressor Animation"
   GraphicView "Graphic view_93" at 838,105 size 48x132; Picture "Graphic_248"
   GraphicView "Graphic view_2" at 823,160 size 19x12; Picture "Graphic_63"
   GraphicView "Graphic view_79" at 823,197 size 19x12; Picture "Graphic_63"
   Bar "Bar_1" at 852,115 size 20x105; Unit  %; MinimumValue 0; MaximumValue 100
      ProcessValue <- "12_AI_Data_PIT112In_SCALED"
      MaximumValue <- "84_Setpoints_PIT112_HighHigh"
   Button "HmiScreenItemData_4" at 1129,1 size 150x43; TextOn 'I&A Compressor Ok'; TextOff 'Back'
      on Release: function_efd93a16()
   IOField "I/O field_20" at 431,212 size 70x25; FormatPattern 99.99; Unit  Bar
      ProcessValue <- "12_AI_Data_PIT112In_SCALED"
   TextField "Text field_28" at 307,216 size 126x18; Text 'System Pressure'
   TextField "Text field_10" at 306,584 size 173x20; Text 'Air / Inert Gas Pressure'
   Button "Button_9" at 630,581 size 57x25; TextOn 'Enabled'; TextOff 'Text'
   TextField "Text field_17" at 306,620 size 310x20; Text 'Air / Inert Gas Pressure Setpoint (Pre-Ignition)'
   Button "Button_11" at 630,618 size 57x25; TextOn 'Enabled'; TextOff 'Text'
   TextField "Text field_12" at 311,736 size 182x20; Text 'Modulating Valve Position'
   TextField "Text field_25" at 306,657 size 310x20; Text 'Air / Inert Gas Pressure Setpoint (Post-Ignition)'
   Button "Button_10" at 630,655 size 57x25; TextOn 'Enabled'; TextOff 'Text'
   IOField "I/O field_2" at 625,582 size 66x25; FormatPattern 999; Unit  mbar
      ProcessValue <- "12_AI_Data_PIT402_SCALED"
   IOField "I/O field_3" at 625,618 size 66x25; Authorization "Commissioning"; FormatPattern 999; Unit  mbar
      ProcessValue <- "84_Setpoints_PIT402_Pilot_Target"
   IOField "I/O field_6" at 625,734 size 66x25; FormatPattern 999; Unit  %
      ProcessValue <- "16_AQ_Data_CV403_CNTRL"
   IOField "I/O field_7" at 625,692 size 66x23; FormatPattern 999; Unit  mBar
      ProcessValue <- "19_AUTO_CMNDS_Data_PIT402_Target"
      Appearance <- "19_AUTO_CMNDS_Data_PIT402_Target"
   IOField "I/O field_12" at 625,655 size 66x25; Authorization "Commissioning"; FormatPattern 999; Unit  mbar